   If SmartTags("SDC\DB_SDC_TS_REFERENCE\_TS_Ref_Nr") >= SmartTags("DB_SDC_TS_REFERENCE_5_HEADER.MIN_NR_SEK") And SmartTags("SDC\DB_SDC_TS_REFERENCE\_TS_Ref_Nr") <= SmartTags("DB_SDC_TS_REFERENCE_5_HEADER.MAX_NR_SEK") Then
   
      SmartTags("SDC\DB_SDC_TS_REFERENCE\_TS_Ref_DB_Nr") = SmartTags("DB_SDC_TS_REFERENCE_5_HEADER.DB_NR")   
   
      TS_Nr = TS_Nr - SmartTags("DB_SDC_TS_REFERENCE_5_HEADER.MIN_NR_SEK") + 1
   
      SmartTags("SDC\DB_SDC_TS_REFERENCE\_TS_Ref_Byte_00")  =   0 + TS_Nr * Laenge_Data - Laenge_Data + Allg_Offset
      SmartTags("SDC\DB_SDC_TS_REFERENCE\_TS_Ref_Byte_16")  =  16 + TS_Nr * Laenge_Data - Laenge_Data + Allg_Offset  
      SmartTags("SDC\DB_SDC_TS_REFERENCE\_TS_Ref_Byte_32")  =  32 + TS_Nr * Laenge_Data - Laenge_Data + Allg_Offset  
      SmartTags("SDC\DB_SDC_TS_REFERENCE\_TS_Ref_Byte_48")  =  48 + TS_Nr * Laenge_Data - Laenge_Data + Allg_Offset   
      SmartTags("SDC\DB_SDC_TS_REFERENCE\_TS_Ref_Byte_64")  =  64 + TS_Nr * Laenge_Data - Laenge_Data + Allg_Offset   
      SmartTags("SDC\DB_SDC_TS_REFERENCE\_TS_Ref_Byte_80")  =  80 + TS_Nr * Laenge_Data - Laenge_Data + Allg_Offset   
      SmartTags("SDC\DB_SDC_TS_REFERENCE\_TS_Ref_Byte_96")  =  96 + TS_Nr * Laenge_Data - Laenge_Data + Allg_Offset 
      SmartTags("SDC\DB_SDC_TS_REFERENCE\_TS_Ref_Byte_112") = 112 + TS_Nr * Laenge_Data - Laenge_Data + Allg_Offset      
    
   End If
   
   If SmartTags("SDC\DB_SDC_TS_REFERENCE\_TS_Ref_Nr") >= SmartTags("DB_SDC_TS_REFERENCE_6_HEADER.MIN_NR_SEK") And SmartTags("SDC\DB_SDC_TS_REFERENCE\_TS_Ref_Nr") <= SmartTags("DB_SDC_TS_REFERENCE_6_HEADER.MAX_NR_SEK") Then
   
      SmartTags("SDC\DB_SDC_TS_REFERENCE\_TS_Ref_DB_Nr") = SmartTags("DB_SDC_TS_REFERENCE_6_HEADER.DB_NR")   
   
      TS_Nr = TS_Nr - SmartTags("DB_SDC_TS_REFERENCE_6_HEADER.MIN_NR_SEK") + 1
   
      SmartTags("SDC\DB_SDC_TS_REFERENCE\_TS_Ref_Byte_00")  =   0 + TS_Nr * Laenge_Data - Laenge_Data + Allg_Offset
      SmartTags("SDC\DB_SDC_TS_REFERENCE\_TS_Ref_Byte_16")  =  16 + TS_Nr * Laenge_Data - Laenge_Data + Allg_Offset  
      SmartTags("SDC\DB_SDC_TS_REFERENCE\_TS_Ref_Byte_32")  =  32 + TS_Nr * Laenge_Data - Laenge_Data + Allg_Offset  
      SmartTags("SDC\DB_SDC_TS_REFERENCE\_TS_Ref_Byte_48")  =  48 + TS_Nr * Laenge_Data - Laenge_Data + Allg_Offset   
      SmartTags("SDC\DB_SDC_TS_REFERENCE\_TS_Ref_Byte_64")  =  64 + TS_Nr * Laenge_Data - Laenge_Data + Allg_Offset   
      SmartTags("SDC\DB_SDC_TS_REFERENCE\_TS_Ref_Byte_80")  =  80 + TS_Nr * Laenge_Data - Laenge_Data + Allg_Offset   
      SmartTags("SDC\DB_SDC_TS_REFERENCE\_TS_Ref_Byte_96")  =  96 + TS_Nr * Laenge_Data - Laenge_Data + Allg_Offset 
      SmartTags("SDC\DB_SDC_TS_REFERENCE\_TS_Ref_Byte_112") = 112 + TS_Nr * Laenge_Data - Laenge_Data + Allg_Offset      
     
   End If   

VB script "SDC_INIT"
   'Tip:
   ' 1. Verwenden Sie die Tastenkombination <CTRL+SPACE> oder <CTRL+I>, um eine Liste aller Objekte und Funktionen zu öffnen
   ' 2. Schreiben Sie den Code unter Verwendung des HMI Runtime Objekts.
   '  Beispiel: HmiRuntime.Screens("Screen_1").
   ' 3. Verwenden Sie die Tastenkombination <CTRL+J>, um eine Objektreferenz zu erstellen.
   'Schreiben Sie den Code ab dieser Position:
   
    SmartTags("_intern_Pult_Nr") = 21 ' SmartTags("__DB_Pult") - 209

VB script "SDC_FILL_intNR"
   'Tip:
   ' 1. Verwenden Sie die Tastenkombination <CTRL+SPACE> oder <CTRL+I>, um eine Liste aller Objekte und Funktionen zu öffnen
   ' 2. Schreiben Sie den Code unter Verwendung des HMI Runtime Objekts.
   '  Beispiel: HmiRuntime.Screens("Screen_1").
   ' 3. Verwenden Sie die Tastenkombination <CTRL+J>, um eine Objektreferenz zu erstellen.
   'Schreiben Sie den Code ab dieser Position:
   Dim i
   
   For i=1 To 200 
   	SmartTags("_intern_" & i) = i
   Next
   		

VB script "DecActScreenDev"
     If (SmartTags("UserDiag_HmiData_actScreenDevices") > 1) Then
     	SmartTags("UserDiag_HmiData_actScreenDevices") = SmartTags("UserDiag_HmiData_actScreenDevices") - 1
     End If
     

VB script "IncActScreenDev"
     If (SmartTags("UserDiag_HmiData_actScreenDevices") < SmartTags("UserDiag_HmiData_maxScreensDevices")) Then
     	SmartTags("UserDiag_HmiData_actScreenDevices") = SmartTags("UserDiag_HmiData_actScreenDevices") + 1
     End If
     

scheduled task "Reset"
   on Action: SetTag("SDC\_EDIT", 0)
*)

(* ===== HMI "HMI_RT_1" =====

ScreenModuleEditorView "typeDevice" 640x480
   Button "Schaltfläche_3" at 90,10 size 110x110; TextOff 'Text'
      Visibility <- "DeviceNumber"
   Rectangle "Rectangle_1" at 90,10 size 110x110
      Visibility <- "DeviceNumber"
      Appearance <- "ErrorState"
   IOField "EA-Feld_1" at 90,10 size 110x110; FormatPattern 999
      ProcessValue <- "DeviceNumber"
      Visibility <- "DeviceNumber"
*)

(* ===== HMI "HMI_RT_1" =====

ScreenModuleEditorView "typeDevice" 640x480
   Button "Schaltfläche_3" at 90,10 size 110x65; TextOff 'Text'
      Visibility <- "DeviceNumber"
   Rectangle "Rectangle_1" at 90,10 size 110x65
      Visibility <- "DeviceNumber"
      Appearance <- "ErrorState"
   IOField "EA-Feld_1" at 90,10 size 110x65; FormatPattern 999
      Visibility <- "DeviceNumber"
      ProcessValue <- "DeviceNumber"
*)